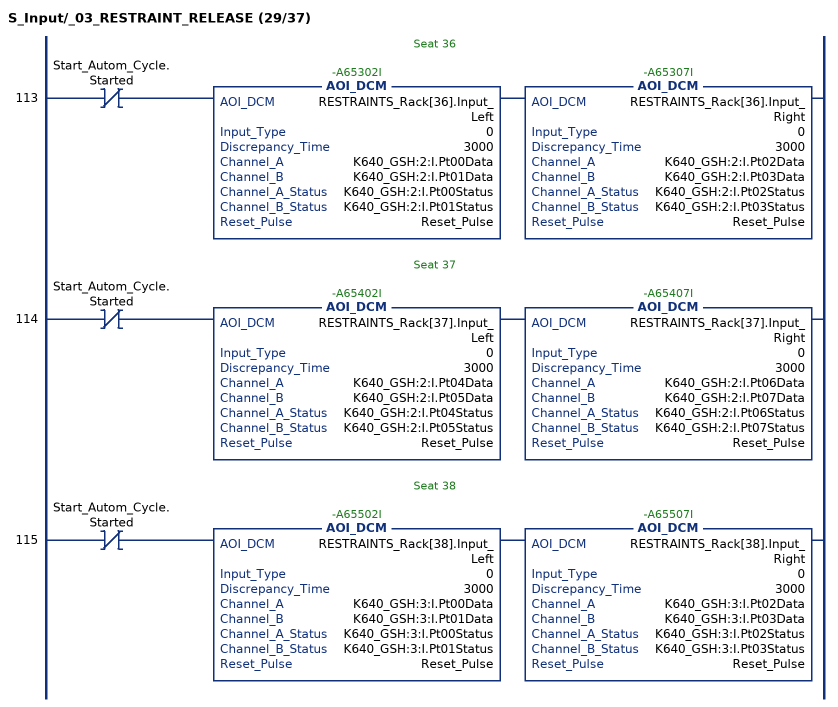
   // Seat 36
   113: XIO(Start_Autom_Cycle.Started)AOI_DCM(RESTRAINTS_Rack[36].Input_Left,0,3000,K640_GSH:2:I.Pt00Data,K640_GSH:2:I.Pt01Data,K640_GSH:2:I.Pt00Status,K640_GSH:2:I.Pt01Status,Reset_Pulse)AOI_DCM(RESTRAINTS_Rack[36].Input_Right,0,3000,K640_GSH:2:I.Pt02Data,K640_GSH:2:I.Pt03Data,K640_GSH:2:I.Pt02Status,K640_GSH:2:I.Pt03Status,Reset_Pulse);
   // Seat 37
   114: XIO(Start_Autom_Cycle.Started)AOI_DCM(RESTRAINTS_Rack[37].Input_Left,0,3000,K640_GSH:2:I.Pt04Data,K640_GSH:2:I.Pt05Data,K640_GSH:2:I.Pt04Status,K640_GSH:2:I.Pt05Status,Reset_Pulse)AOI_DCM(RESTRAINTS_Rack[37].Input_Right,0,3000,K640_GSH:2:I.Pt06Data,K640_GSH:2:I.Pt07Data,K640_GSH:2:I.Pt06Status,K640_GSH:2:I.Pt07Status,Reset_Pulse);
   // Seat 38
   115: XIO(Start_Autom_Cycle.Started)AOI_DCM(RESTRAINTS_Rack[38].Input_Left,0,3000,K640_GSH:3:I.Pt00Data,K640_GSH:3:I.Pt01Data,K640_GSH:3:I.Pt00Status,K640_GSH:3:I.Pt01Status,Reset_Pulse)AOI_DCM(RESTRAINTS_Rack[38].Input_Right,0,3000,K640_GSH:3:I.Pt02Data,K640_GSH:3:I.Pt03Data,K640_GSH:3:I.Pt02Status,K640_GSH:3:I.Pt03Status,Reset_Pulse);
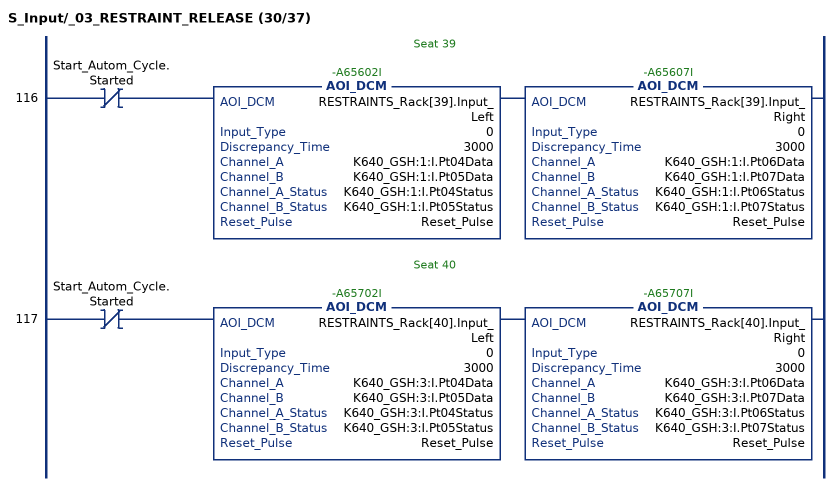
   // Seat 39
   116: XIO(Start_Autom_Cycle.Started)AOI_DCM(RESTRAINTS_Rack[39].Input_Left,0,3000,K640_GSH:1:I.Pt04Data,K640_GSH:1:I.Pt05Data,K640_GSH:1:I.Pt04Status,K640_GSH:1:I.Pt05Status,Reset_Pulse)AOI_DCM(RESTRAINTS_Rack[39].Input_Right,0,3000,K640_GSH:1:I.Pt06Data,K640_GSH:1:I.Pt07Data,K640_GSH:1:I.Pt06Status,K640_GSH:1:I.Pt07Status,Reset_Pulse);
   // Seat 40
   117: XIO(Start_Autom_Cycle.Started)AOI_DCM(RESTRAINTS_Rack[40].Input_Left,0,3000,K640_GSH:3:I.Pt04Data,K640_GSH:3:I.Pt05Data,K640_GSH:3:I.Pt04Status,K640_GSH:3:I.Pt05Status,Reset_Pulse)AOI_DCM(RESTRAINTS_Rack[40].Input_Right,0,3000,K640_GSH:3:I.Pt06Data,K640_GSH:3:I.Pt07Data,K640_GSH:3:I.Pt06Status,K640_GSH:3:I.Pt07Status,Reset_Pulse);
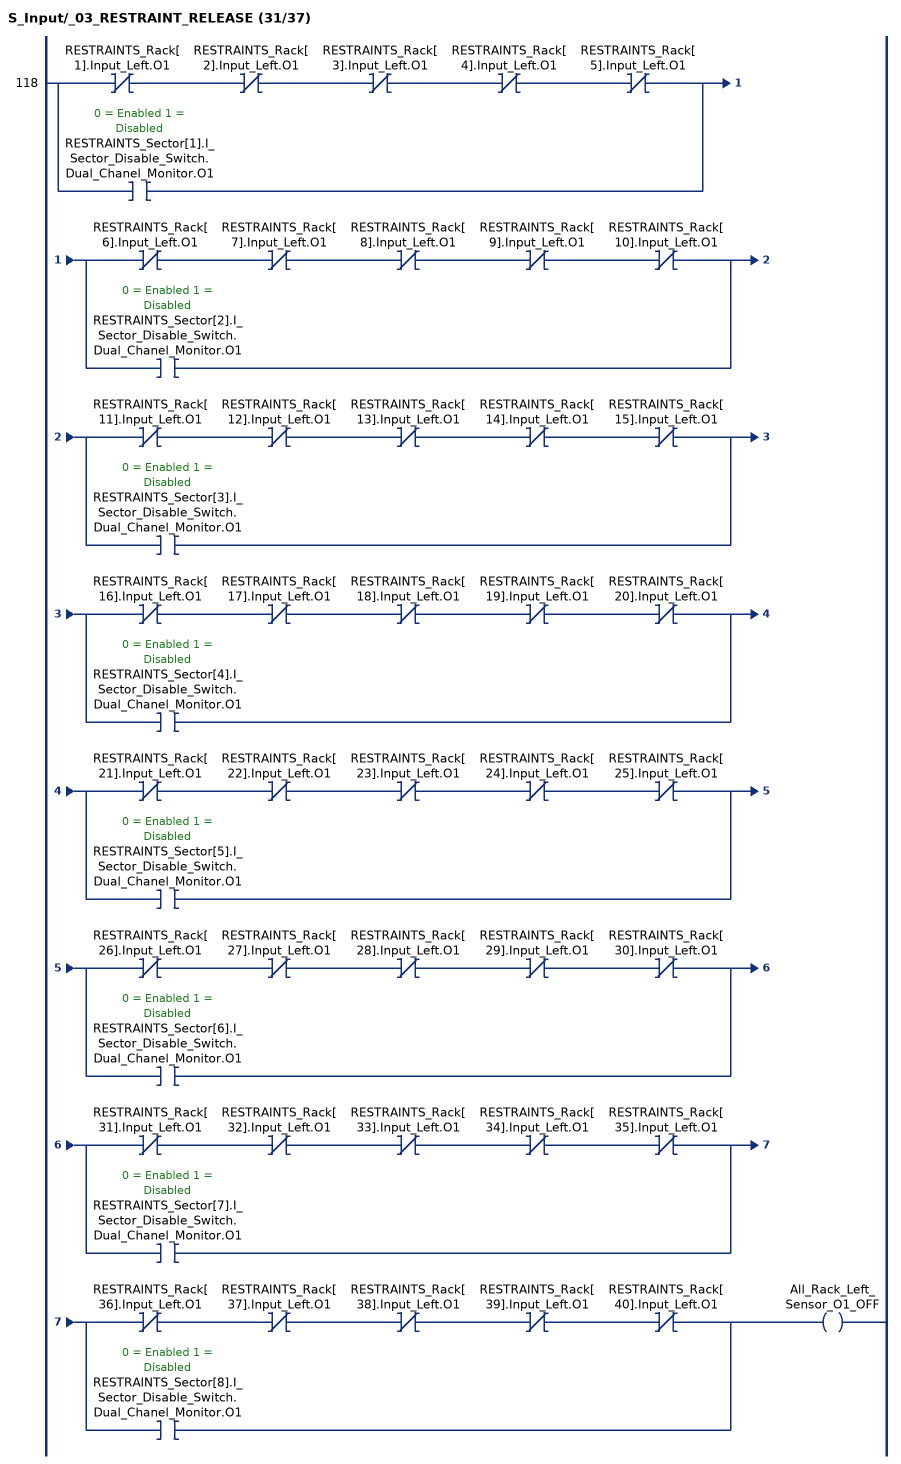
   118: [XIO(RESTRAINTS_Rack[1].Input_Left.O1) XIO(RESTRAINTS_Rack[2].Input_Left.O1) XIO(RESTRAINTS_Rack[3].Input_Left.O1) XIO(RESTRAINTS_Rack[4].Input_Left.O1) XIO(RESTRAINTS_Rack[5].Input_Left.O1) ,XIC(RESTRAINTS_Sector[1].I_Sector_Disable_Switch.Dual_Chanel_Monitor.O1) ][XIO(RESTRAINTS_Rack[6].Input_Left.O1) XIO(RESTRAINTS_Rack[7].Input_Left.O1) XIO(RESTRAINTS_Rack[8].Input_Left.O1) XIO(RESTRAINTS_Rack[9].Input_Left.O1) XIO(RESTRAINTS_Rack[10].Input_Left.O1) ,XIC(RESTRAINTS_Sector[2].I_Sector_Disable_Switch.Dual_Chanel_Monitor.O1) ][XIO(RESTRAINTS_Rack[11].Input_Left.O1) XIO(RESTRAINTS_Rack[12].Input_Left.O1) XIO(RESTRAINTS_Rack[13].Input_Left.O1) XIO(RESTRAINTS_Rack[14].Input_Left.O1) XIO(RESTRAINTS_Rack[15].Input_Left.O1) ,XIC(RESTRAINTS_Sector[3].I_Sector_Disable_Switch.Dual_Chanel_Monitor.O1) ][XIO(RESTRAINTS_Rack[16].Input_Left.O1) XIO(RESTRAINTS_Rack[17].Input_Left.O1) XIO(RESTRAINTS_Rack[18].Input_Left.O1) XIO(RESTRAINTS_Rack[19].Input_Left.O1) XIO(RESTRAINTS_Rack[20].Input_Left.O1) ,XIC(RESTRAINTS_Sector[4].I_Sector_Disable_Switch.Dual_Chanel_Monitor.O1) ][XIO(RESTRAINTS_Rack[21].Input_Left.O1) XIO(RESTRAINTS_Rack[22].Input_Left.O1) XIO(RESTRAINTS_Rack[23].Input_Left.O1) XIO(RESTRAINTS_Rack[24].Input_Left.O1) XIO(RESTRAINTS_Rack[25].Input_Left.O1) ,XIC(RESTRAINTS_Sector[5].I_Sector_Disable_Switch.Dual_Chanel_Monitor.O1) ][XIO(RESTRAINTS_Rack[26].Input_Left.O1) XIO(RESTRAINTS_Rack[27].Input_Left.O1) XIO(RESTRAINTS_Rack[28].Input_Left.O1) XIO(RESTRAINTS_Rack[29].Input_Left.O1) XIO(RESTRAINTS_Rack[30].Input_Left.O1) ,XIC(RESTRAINTS_Sector[6].I_Sector_Disable_Switch.Dual_Chanel_Monitor.O1) ][XIO(RESTRAINTS_Rack[31].Input_Left.O1) XIO(RESTRAINTS_Rack[32].Input_Left.O1) XIO(RESTRAINTS_Rack[33].Input_Left.O1) XIO(RESTRAINTS_Rack[34].Input_Left.O1) XIO(RESTRAINTS_Rack[35].Input_Left.O1) ,XIC(RESTRAINTS_Sector[7].I_Sector_Disable_Switch.Dual_Chanel_Monitor.O1) ][XIO(RESTRAINTS_Rack[36].Input_Left.O1) XIO(RESTRAINTS_Rack[37].Input_Left.O1) XIO(RESTRAINTS_Rack[38].Input_Left.O1) XIO(RESTRAINTS_Rack[39].Input_Left.O1) XIO(RESTRAINTS_Rack[40].Input_Left.O1) ,XIC(RESTRAINTS_Sector[8].I_Sector_Disable_Switch.Dual_Chanel_Monitor.O1) ]OTE(All_Rack_Left_Sensor_O1_OFF);
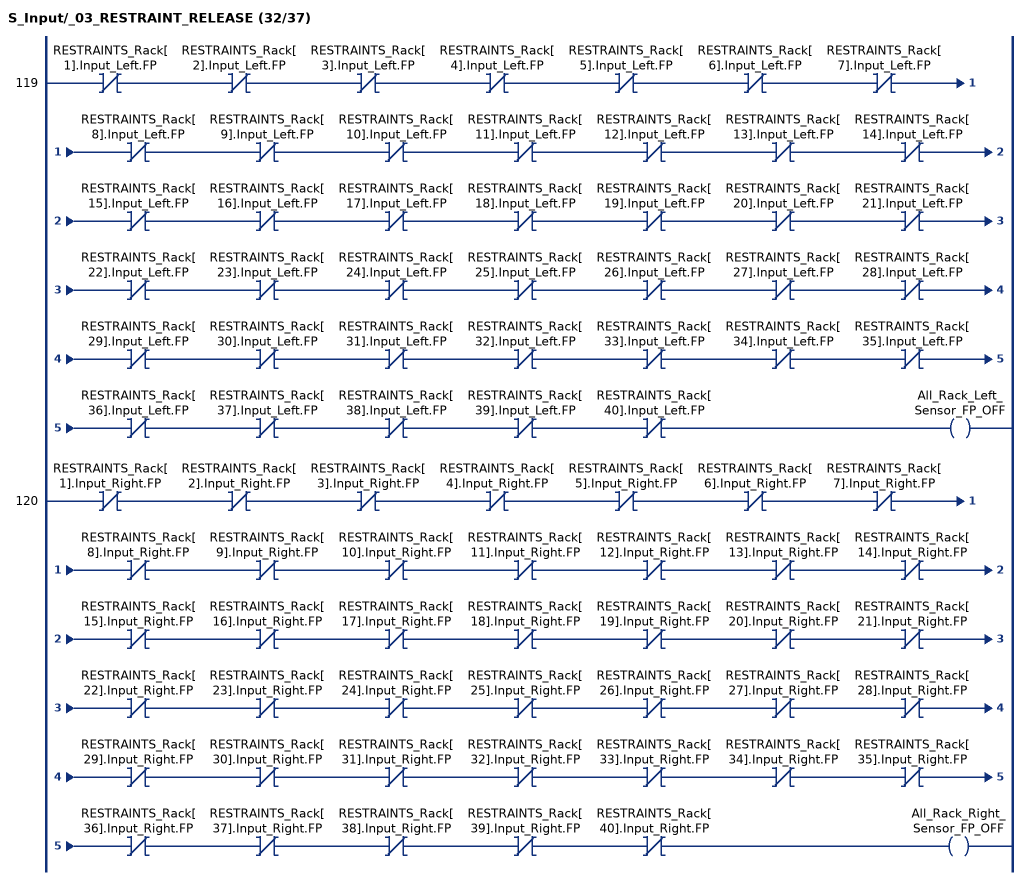
   119: XIO(RESTRAINTS_Rack[1].Input_Left.FP)XIO(RESTRAINTS_Rack[2].Input_Left.FP)XIO(RESTRAINTS_Rack[3].Input_Left.FP)XIO(RESTRAINTS_Rack[4].Input_Left.FP)XIO(RESTRAINTS_Rack[5].Input_Left.FP)XIO(RESTRAINTS_Rack[6].Input_Left.FP)XIO(RESTRAINTS_Rack[7].Input_Left.FP)XIO(RESTRAINTS_Rack[8].Input_Left.FP)XIO(RESTRAINTS_Rack[9].Input_Left.FP)XIO(RESTRAINTS_Rack[10].Input_Left.FP)XIO(RESTRAINTS_Rack[11].Input_Left.FP)XIO(RESTRAINTS_Rack[12].Input_Left.FP)XIO(RESTRAINTS_Rack[13].Input_Left.FP)XIO(RESTRAINTS_Rack[14].Input_Left.FP)XIO(RESTRAINTS_Rack[15].Input_Left.FP)XIO(RESTRAINTS_Rack[16].Input_Left.FP)XIO(RESTRAINTS_Rack[17].Input_Left.FP)XIO(RESTRAINTS_Rack[18].Input_Left.FP)XIO(RESTRAINTS_Rack[19].Input_Left.FP)XIO(RESTRAINTS_Rack[20].Input_Left.FP)XIO(RESTRAINTS_Rack[21].Input_Left.FP)XIO(RESTRAINTS_Rack[22].Input_Left.FP)XIO(RESTRAINTS_Rack[23].Input_Left.FP)XIO(RESTRAINTS_Rack[24].Input_Left.FP)XIO(RESTRAINTS_Rack[25].Input_Left.FP)XIO(RESTRAINTS_Rack[26].Input_Left.FP)XIO(RESTRAINTS_Rack[27].Input_Left.FP)XIO(RESTRAINTS_Rack[28].Input_Left.FP)XIO(RESTRAINTS_Rack[29].Input_Left.FP)XIO(RESTRAINTS_Rack[30].Input_Left.FP)XIO(RESTRAINTS_Rack[31].Input_Left.FP)XIO(RESTRAINTS_Rack[32].Input_Left.FP)XIO(RESTRAINTS_Rack[33].Input_Left.FP)XIO(RESTRAINTS_Rack[34].Input_Left.FP)XIO(RESTRAINTS_Rack[35].Input_Left.FP)XIO(RESTRAINTS_Rack[36].Input_Left.FP)XIO(RESTRAINTS_Rack[37].Input_Left.FP)XIO(RESTRAINTS_Rack[38].Input_Left.FP)XIO(RESTRAINTS_Rack[39].Input_Left.FP)XIO(RESTRAINTS_Rack[40].Input_Left.FP)OTE(All_Rack_Left_Sensor_FP_OFF);
   120: XIO(RESTRAINTS_Rack[1].Input_Right.FP)XIO(RESTRAINTS_Rack[2].Input_Right.FP)XIO(RESTRAINTS_Rack[3].Input_Right.FP)XIO(RESTRAINTS_Rack[4].Input_Right.FP)XIO(RESTRAINTS_Rack[5].Input_Right.FP)XIO(RESTRAINTS_Rack[6].Input_Right.FP)XIO(RESTRAINTS_Rack[7].Input_Right.FP)XIO(RESTRAINTS_Rack[8].Input_Right.FP)XIO(RESTRAINTS_Rack[9].Input_Right.FP)XIO(RESTRAINTS_Rack[10].Input_Right.FP)XIO(RESTRAINTS_Rack[11].Input_Right.FP)XIO(RESTRAINTS_Rack[12].Input_Right.FP)XIO(RESTRAINTS_Rack[13].Input_Right.FP)XIO(RESTRAINTS_Rack[14].Input_Right.FP)XIO(RESTRAINTS_Rack[15].Input_Right.FP)XIO(RESTRAINTS_Rack[16].Input_Right.FP)XIO(RESTRAINTS_Rack[17].Input_Right.FP)XIO(RESTRAINTS_Rack[18].Input_Right.FP)XIO(RESTRAINTS_Rack[19].Input_Right.FP)XIO(RESTRAINTS_Rack[20].Input_Right.FP)XIO(RESTRAINTS_Rack[21].Input_Right.FP)XIO(RESTRAINTS_Rack[22].Input_Right.FP)XIO(RESTRAINTS_Rack[23].Input_Right.FP)XIO(RESTRAINTS_Rack[24].Input_Right.FP)XIO(RESTRAINTS_Rack[25].Input_Right.FP)XIO(RESTRAINTS_Rack[26].Input_Right.FP)XIO(RESTRAINTS_Rack[27].Input_Right.FP)XIO(RESTRAINTS_Rack[28].Input_Right.FP)XIO(RESTRAINTS_Rack[29].Input_Right.FP)XIO(RESTRAINTS_Rack[30].Input_Right.FP)XIO(RESTRAINTS_Rack[31].Input_Right.FP)XIO(RESTRAINTS_Rack[32].Input_Right.FP)XIO(RESTRAINTS_Rack[33].Input_Right.FP)XIO(RESTRAINTS_Rack[34].Input_Right.FP)XIO(RESTRAINTS_Rack[35].Input_Right.FP)XIO(RESTRAINTS_Rack[36].Input_Right.FP)XIO(RESTRAINTS_Rack[37].Input_Right.FP)XIO(RESTRAINTS_Rack[38].Input_Right.FP)XIO(RESTRAINTS_Rack[39].Input_Right.FP)XIO(RESTRAINTS_Rack[40].Input_Right.FP)OTE(All_Rack_Right_Sensor_FP_OFF);
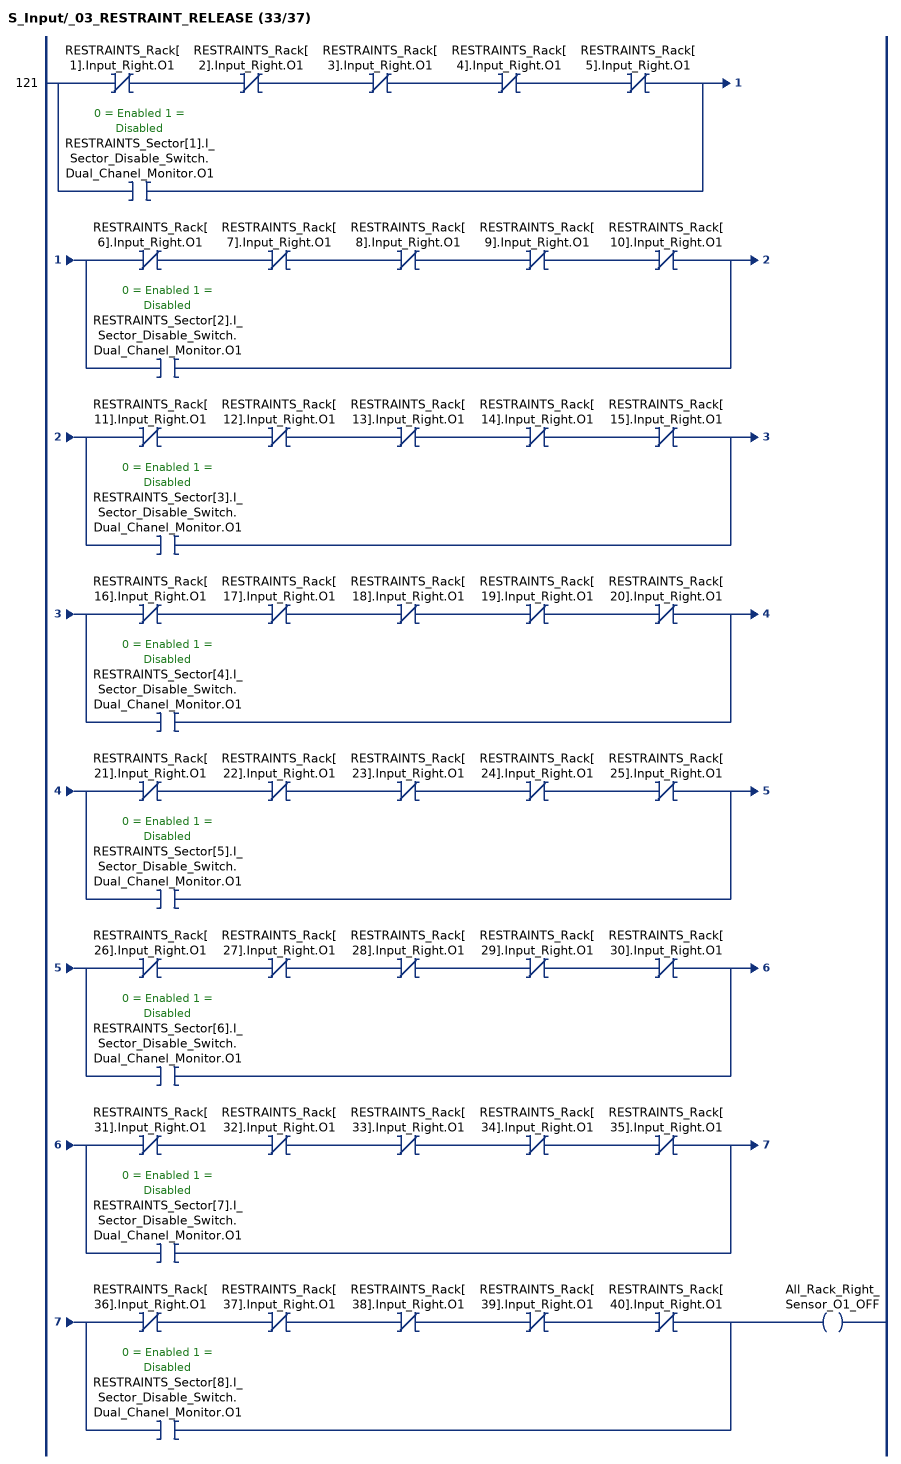
   121: [XIO(RESTRAINTS_Rack[1].Input_Right.O1) XIO(RESTRAINTS_Rack[2].Input_Right.O1) XIO(RESTRAINTS_Rack[3].Input_Right.O1) XIO(RESTRAINTS_Rack[4].Input_Right.O1) XIO(RESTRAINTS_Rack[5].Input_Right.O1) ,XIC(RESTRAINTS_Sector[1].I_Sector_Disable_Switch.Dual_Chanel_Monitor.O1) ][XIO(RESTRAINTS_Rack[6].Input_Right.O1) XIO(RESTRAINTS_Rack[7].Input_Right.O1) XIO(RESTRAINTS_Rack[8].Input_Right.O1) XIO(RESTRAINTS_Rack[9].Input_Right.O1) XIO(RESTRAINTS_Rack[10].Input_Right.O1) ,XIC(RESTRAINTS_Sector[2].I_Sector_Disable_Switch.Dual_Chanel_Monitor.O1) ][XIO(RESTRAINTS_Rack[11].Input_Right.O1) XIO(RESTRAINTS_Rack[12].Input_Right.O1) XIO(RESTRAINTS_Rack[13].Input_Right.O1) XIO(RESTRAINTS_Rack[14].Input_Right.O1) XIO(RESTRAINTS_Rack[15].Input_Right.O1) ,XIC(RESTRAINTS_Sector[3].I_Sector_Disable_Switch.Dual_Chanel_Monitor.O1) ][XIO(RESTRAINTS_Rack[16].Input_Right.O1) XIO(RESTRAINTS_Rack[17].Input_Right.O1) XIO(RESTRAINTS_Rack[18].Input_Right.O1) XIO(RESTRAINTS_Rack[19].Input_Right.O1) XIO(RESTRAINTS_Rack[20].Input_Right.O1) ,XIC(RESTRAINTS_Sector[4].I_Sector_Disable_Switch.Dual_Chanel_Monitor.O1) ][XIO(RESTRAINTS_Rack[21].Input_Right.O1) XIO(RESTRAINTS_Rack[22].Input_Right.O1) XIO(RESTRAINTS_Rack[23].Input_Right.O1) XIO(RESTRAINTS_Rack[24].Input_Right.O1) XIO(RESTRAINTS_Rack[25].Input_Right.O1) ,XIC(RESTRAINTS_Sector[5].I_Sector_Disable_Switch.Dual_Chanel_Monitor.O1) ][XIO(RESTRAINTS_Rack[26].Input_Right.O1) XIO(RESTRAINTS_Rack[27].Input_Right.O1) XIO(RESTRAINTS_Rack[28].Input_Right.O1) XIO(RESTRAINTS_Rack[29].Input_Right.O1) XIO(RESTRAINTS_Rack[30].Input_Right.O1) ,XIC(RESTRAINTS_Sector[6].I_Sector_Disable_Switch.Dual_Chanel_Monitor.O1) ][XIO(RESTRAINTS_Rack[31].Input_Right.O1) XIO(RESTRAINTS_Rack[32].Input_Right.O1) XIO(RESTRAINTS_Rack[33].Input_Right.O1) XIO(RESTRAINTS_Rack[34].Input_Right.O1) XIO(RESTRAINTS_Rack[35].Input_Right.O1) ,XIC(RESTRAINTS_Sector[7].I_Sector_Disable_Switch.Dual_Chanel_Monitor.O1) ][XIO(RESTRAINTS_Rack[36].Input_Right.O1) XIO(RESTRAINTS_Rack[37].Input_Right.O1) XIO(RESTRAINTS_Rack[38].Input_Right.O1) XIO(RESTRAINTS_Rack[39].Input_Right.O1) XIO(RESTRAINTS_Rack[40].Input_Right.O1) ,XIC(RESTRAINTS_Sector[8].I_Sector_Disable_Switch.Dual_Chanel_Monitor.O1) ]OTE(All_Rack_Right_Sensor_O1_OFF);
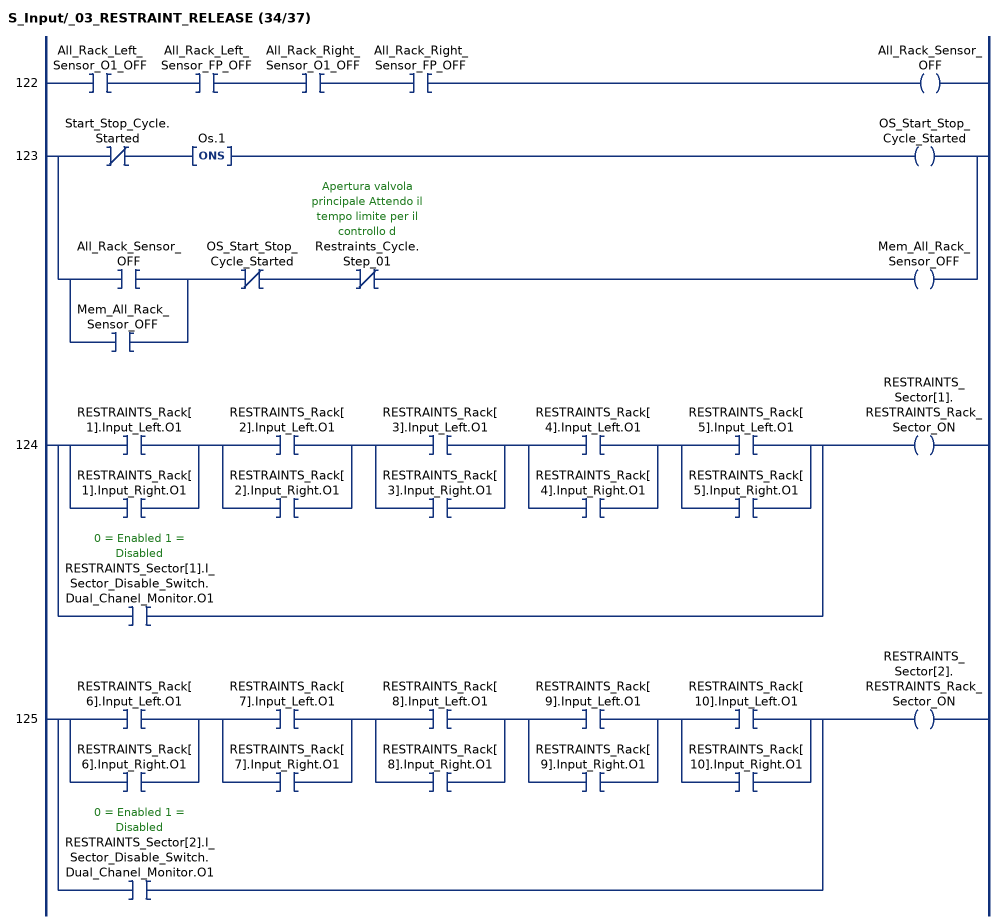
   122: XIC(All_Rack_Left_Sensor_O1_OFF)XIC(All_Rack_Left_Sensor_FP_OFF)XIC(All_Rack_Right_Sensor_O1_OFF)XIC(All_Rack_Right_Sensor_FP_OFF)OTE(All_Rack_Sensor_OFF);
   123: [XIO(Start_Stop_Cycle.Started) ONS(Os.1) OTE(OS_Start_Stop_Cycle_Started) ,[XIC(All_Rack_Sensor_OFF) ,XIC(Mem_All_Rack_Sensor_OFF) ] XIO(OS_Start_Stop_Cycle_Started) XIO(Restraints_Cycle.Step_01) OTE(Mem_All_Rack_Sensor_OFF) ];
   124: [[XIC(RESTRAINTS_Rack[1].Input_Left.O1) ,XIC(RESTRAINTS_Rack[1].Input_Right.O1) ] [XIC(RESTRAINTS_Rack[2].Input_Left.O1) ,XIC(RESTRAINTS_Rack[2].Input_Right.O1) ] [XIC(RESTRAINTS_Rack[3].Input_Left.O1) ,XIC(RESTRAINTS_Rack[3].Input_Right.O1) ] [XIC(RESTRAINTS_Rack[4].Input_Left.O1) ,XIC(RESTRAINTS_Rack[4].Input_Right.O1) ] [XIC(RESTRAINTS_Rack[5].Input_Left.O1) ,XIC(RESTRAINTS_Rack[5].Input_Right.O1) ] ,XIC(RESTRAINTS_Sector[1].I_Sector_Disable_Switch.Dual_Chanel_Monitor.O1) ]OTE(RESTRAINTS_Sector[1].RESTRAINTS_Rack_Sector_ON);
   125: [[XIC(RESTRAINTS_Rack[6].Input_Left.O1) ,XIC(RESTRAINTS_Rack[6].Input_Right.O1) ] [XIC(RESTRAINTS_Rack[7].Input_Left.O1) ,XIC(RESTRAINTS_Rack[7].Input_Right.O1) ] [XIC(RESTRAINTS_Rack[8].Input_Left.O1) ,XIC(RESTRAINTS_Rack[8].Input_Right.O1) ] [XIC(RESTRAINTS_Rack[9].Input_Left.O1) ,XIC(RESTRAINTS_Rack[9].Input_Right.O1) ] [XIC(RESTRAINTS_Rack[10].Input_Left.O1) ,XIC(RESTRAINTS_Rack[10].Input_Right.O1) ] ,XIC(RESTRAINTS_Sector[2].I_Sector_Disable_Switch.Dual_Chanel_Monitor.O1) ]OTE(RESTRAINTS_Sector[2].RESTRAINTS_Rack_Sector_ON);
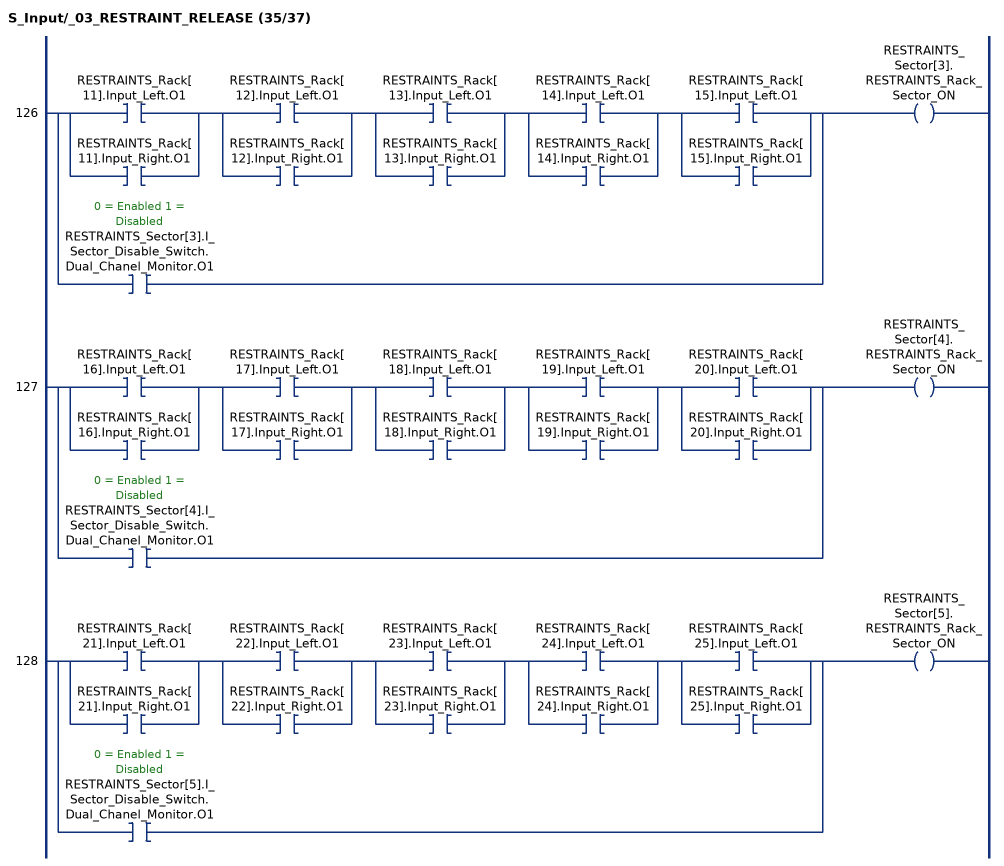
   126: [[XIC(RESTRAINTS_Rack[11].Input_Left.O1) ,XIC(RESTRAINTS_Rack[11].Input_Right.O1) ] [XIC(RESTRAINTS_Rack[12].Input_Left.O1) ,XIC(RESTRAINTS_Rack[12].Input_Right.O1) ] [XIC(RESTRAINTS_Rack[13].Input_Left.O1) ,XIC(RESTRAINTS_Rack[13].Input_Right.O1) ] [XIC(RESTRAINTS_Rack[14].Input_Left.O1) ,XIC(RESTRAINTS_Rack[14].Input_Right.O1) ] [XIC(RESTRAINTS_Rack[15].Input_Left.O1) ,XIC(RESTRAINTS_Rack[15].Input_Right.O1) ] ,XIC(RESTRAINTS_Sector[3].I_Sector_Disable_Switch.Dual_Chanel_Monitor.O1) ]OTE(RESTRAINTS_Sector[3].RESTRAINTS_Rack_Sector_ON);
   127: [[XIC(RESTRAINTS_Rack[16].Input_Left.O1) ,XIC(RESTRAINTS_Rack[16].Input_Right.O1) ] [XIC(RESTRAINTS_Rack[17].Input_Left.O1) ,XIC(RESTRAINTS_Rack[17].Input_Right.O1) ] [XIC(RESTRAINTS_Rack[18].Input_Left.O1) ,XIC(RESTRAINTS_Rack[18].Input_Right.O1) ] [XIC(RESTRAINTS_Rack[19].Input_Left.O1) ,XIC(RESTRAINTS_Rack[19].Input_Right.O1) ] [XIC(RESTRAINTS_Rack[20].Input_Left.O1) ,XIC(RESTRAINTS_Rack[20].Input_Right.O1) ] ,XIC(RESTRAINTS_Sector[4].I_Sector_Disable_Switch.Dual_Chanel_Monitor.O1) ]OTE(RESTRAINTS_Sector[4].RESTRAINTS_Rack_Sector_ON);
   128: [[XIC(RESTRAINTS_Rack[21].Input_Left.O1) ,XIC(RESTRAINTS_Rack[21].Input_Right.O1) ] [XIC(RESTRAINTS_Rack[22].Input_Left.O1) ,XIC(RESTRAINTS_Rack[22].Input_Right.O1) ] [XIC(RESTRAINTS_Rack[23].Input_Left.O1) ,XIC(RESTRAINTS_Rack[23].Input_Right.O1) ] [XIC(RESTRAINTS_Rack[24].Input_Left.O1) ,XIC(RESTRAINTS_Rack[24].Input_Right.O1) ] [XIC(RESTRAINTS_Rack[25].Input_Left.O1) ,XIC(RESTRAINTS_Rack[25].Input_Right.O1) ] ,XIC(RESTRAINTS_Sector[5].I_Sector_Disable_Switch.Dual_Chanel_Monitor.O1) ]OTE(RESTRAINTS_Sector[5].RESTRAINTS_Rack_Sector_ON);
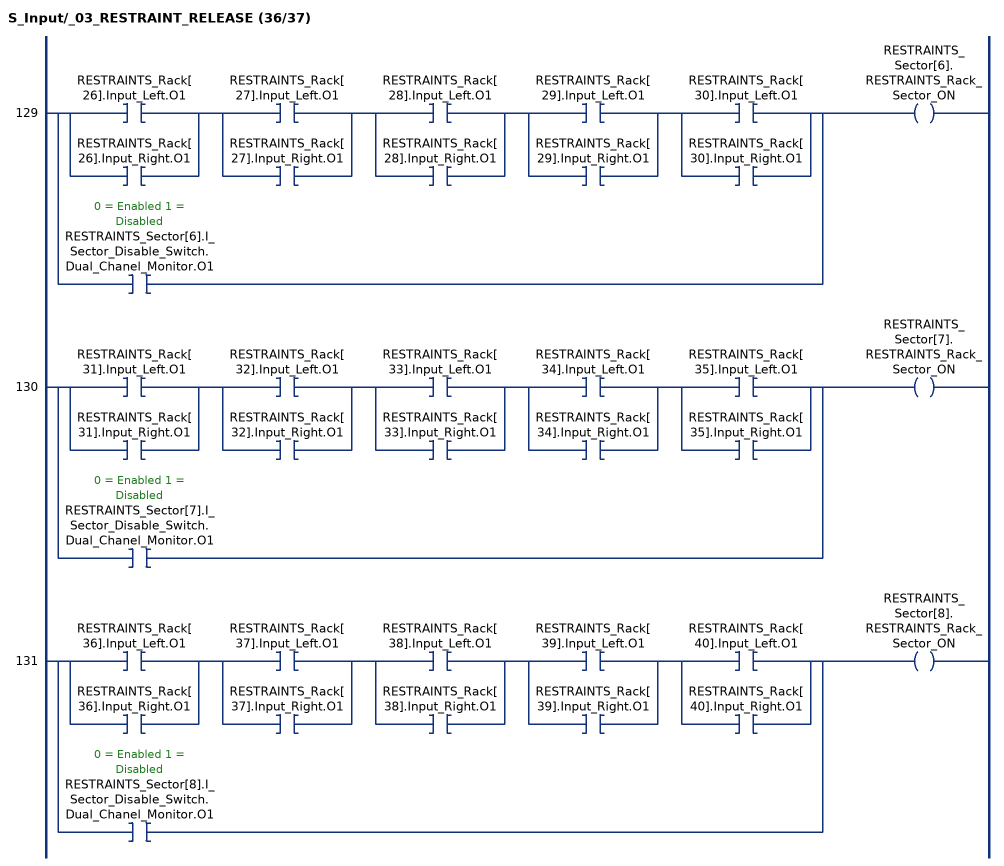
   129: [[XIC(RESTRAINTS_Rack[26].Input_Left.O1) ,XIC(RESTRAINTS_Rack[26].Input_Right.O1) ] [XIC(RESTRAINTS_Rack[27].Input_Left.O1) ,XIC(RESTRAINTS_Rack[27].Input_Right.O1) ] [XIC(RESTRAINTS_Rack[28].Input_Left.O1) ,XIC(RESTRAINTS_Rack[28].Input_Right.O1) ] [XIC(RESTRAINTS_Rack[29].Input_Left.O1) ,XIC(RESTRAINTS_Rack[29].Input_Right.O1) ] [XIC(RESTRAINTS_Rack[30].Input_Left.O1) ,XIC(RESTRAINTS_Rack[30].Input_Right.O1) ] ,XIC(RESTRAINTS_Sector[6].I_Sector_Disable_Switch.Dual_Chanel_Monitor.O1) ]OTE(RESTRAINTS_Sector[6].RESTRAINTS_Rack_Sector_ON);
   130: [[XIC(RESTRAINTS_Rack[31].Input_Left.O1) ,XIC(RESTRAINTS_Rack[31].Input_Right.O1) ] [XIC(RESTRAINTS_Rack[32].Input_Left.O1) ,XIC(RESTRAINTS_Rack[32].Input_Right.O1) ] [XIC(RESTRAINTS_Rack[33].Input_Left.O1) ,XIC(RESTRAINTS_Rack[33].Input_Right.O1) ] [XIC(RESTRAINTS_Rack[34].Input_Left.O1) ,XIC(RESTRAINTS_Rack[34].Input_Right.O1) ] [XIC(RESTRAINTS_Rack[35].Input_Left.O1) ,XIC(RESTRAINTS_Rack[35].Input_Right.O1) ] ,XIC(RESTRAINTS_Sector[7].I_Sector_Disable_Switch.Dual_Chanel_Monitor.O1) ]OTE(RESTRAINTS_Sector[7].RESTRAINTS_Rack_Sector_ON);
   131: [[XIC(RESTRAINTS_Rack[36].Input_Left.O1) ,XIC(RESTRAINTS_Rack[36].Input_Right.O1) ] [XIC(RESTRAINTS_Rack[37].Input_Left.O1) ,XIC(RESTRAINTS_Rack[37].Input_Right.O1) ] [XIC(RESTRAINTS_Rack[38].Input_Left.O1) ,XIC(RESTRAINTS_Rack[38].Input_Right.O1) ] [XIC(RESTRAINTS_Rack[39].Input_Left.O1) ,XIC(RESTRAINTS_Rack[39].Input_Right.O1) ] [XIC(RESTRAINTS_Rack[40].Input_Left.O1) ,XIC(RESTRAINTS_Rack[40].Input_Right.O1) ] ,XIC(RESTRAINTS_Sector[8].I_Sector_Disable_Switch.Dual_Chanel_Monitor.O1) ]OTE(RESTRAINTS_Sector[8].RESTRAINTS_Rack_Sector_ON);
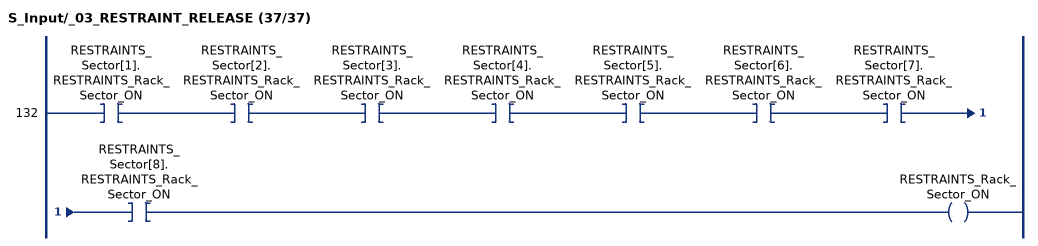
   132: XIC(RESTRAINTS_Sector[1].RESTRAINTS_Rack_Sector_ON)XIC(RESTRAINTS_Sector[2].RESTRAINTS_Rack_Sector_ON)XIC(RESTRAINTS_Sector[3].RESTRAINTS_Rack_Sector_ON)XIC(RESTRAINTS_Sector[4].RESTRAINTS_Rack_Sector_ON)XIC(RESTRAINTS_Sector[5].RESTRAINTS_Rack_Sector_ON)XIC(RESTRAINTS_Sector[6].RESTRAINTS_Rack_Sector_ON)XIC(RESTRAINTS_Sector[7].RESTRAINTS_Rack_Sector_ON)XIC(RESTRAINTS_Sector[8].RESTRAINTS_Rack_Sector_ON)OTE(RESTRAINTS_Rack_Sector_ON);
END_ROUTINE
